   "SDC\DB_SDC_EMS_FLAGS\DB_SDC_EMS_FLAGS.EMS[99]" : Int AT %DB0.DBW0, 1 s
   "SDC\DB_SDC_EMS_FLAGS\DB_SDC_EMS_FLAGS.EMS[100]" : Int AT %DB0.DBW0, 1 s
   "SDC\DB_SDC_EMS_FLAGS\DB_SDC_EMS_FLAGS.EMS[101]" : Int AT %DB0.DBW0, 1 s
   "SDC\DB_SDC_EMS_FLAGS\DB_SDC_EMS_FLAGS.EMS[102]" : Int AT %DB0.DBW0, 1 s
   "SDC\DB_SDC_EMS_FLAGS\DB_SDC_EMS_FLAGS.EMS[103]" : Int AT %DB0.DBW0, 1 s
   "SDC\DB_SDC_EMS_FLAGS\DB_SDC_EMS_FLAGS.EMS[104]" : Int AT %DB0.DBW0, 1 s
   "SDC\DB_SDC_EMS_FLAGS\DB_SDC_EMS_FLAGS.EMS[105]" : Int AT %DB0.DBW0, 1 s
   "SDC\DB_SDC_EMS_FLAGS\DB_SDC_EMS_FLAGS.EMS[106]" : Int AT %DB0.DBW0, 1 s
   "SDC\DB_SDC_EMS_FLAGS\DB_SDC_EMS_FLAGS.EMS[107]" : Int AT %DB0.DBW0, 1 s
   "SDC\DB_SDC_EMS_FLAGS\DB_SDC_EMS_FLAGS.EMS[108]" : Int AT %DB0.DBW0, 1 s
   "SDC\DB_SDC_EMS_FLAGS\DB_SDC_EMS_FLAGS.EMS[109]" : Int AT %DB0.DBW0, 1 s
   "SDC\DB_SDC_EMS_FLAGS\_EMS_Flags_Byte_EMS001" : Int, internal
   "SDC\DB_SDC_EMS_FLAGS\_EMS_Flags_Byte_EMS002" : Int, internal
   "SDC\DB_SDC_EMS_FLAGS\_EMS_Flags_Byte_EMS003" : Int, internal
   "SDC\DB_SDC_EMS_FLAGS\_EMS_Flags_Byte_EMS004" : Int, internal
   "SDC\DB_SDC_EMS_FLAGS\_EMS_Flags_Byte_EMS005" : Int, internal
   "SDC\DB_SDC_EMS_FLAGS\_EMS_Flags_Byte_EMS006" : Int, internal
   "SDC\DB_SDC_EMS_FLAGS\_EMS_Flags_Byte_EMS007" : Int, internal
   "SDC\DB_SDC_EMS_FLAGS\_EMS_Flags_Byte_EMS008" : Int, internal
   "SDC\DB_SDC_EMS_FLAGS\_EMS_Flags_Byte_EMS009" : Int, internal
   "SDC\DB_SDC_EMS_FLAGS\_EMS_Flags_Byte_EMS010" : Int, internal
   "SDC\DB_SDC_EMS_FLAGS\_EMS_Flags_Byte_EMS011" : Int, internal
   "SDC\DB_SDC_EMS_FLAGS\_EMS_Flags_Byte_EMS012" : Int, internal
   "SDC\DB_SDC_EMS_FLAGS\_EMS_Flags_Byte_EMS013" : Int, internal
   "SDC\DB_SDC_EMS_FLAGS\_EMS_Flags_Byte_EMS014" : Int, internal
   "SDC\DB_SDC_EMS_FLAGS\_EMS_Flags_Byte_EMS015" : Int, internal
   "SDC\DB_SDC_EMS_FLAGS\_EMS_Flags_Byte_EMS016" : Int, internal
   "SDC\DB_SDC_EMS_FLAGS\_EMS_Flags_Byte_EMS017" : Int, internal
   "SDC\DB_SDC_EMS_FLAGS\_EMS_Flags_Byte_EMS018" : Int, internal
   "SDC\DB_SDC_EMS_FLAGS\_EMS_Flags_Byte_EMS019" : Int, internal
   "SDC\DB_SDC_EMS_FLAGS\_EMS_Flags_Byte_EMS020" : Int, internal
   "SDC\DB_SDC_EMS_FLAGS\_EMS_Flags_Byte_EMS021" : Int, internal
   "SDC\DB_SDC_EMS_FLAGS\_EMS_Flags_Byte_EMS022" : Int, internal
   "SDC\DB_SDC_EMS_FLAGS\_EMS_Flags_Byte_EMS023" : Int, internal
   "SDC\DB_SDC_EMS_FLAGS\_EMS_Flags_Byte_EMS024" : Int, internal
   "SDC\DB_SDC_EMS_FLAGS\_EMS_Flags_Byte_EMS025" : Int, internal
   "SDC\DB_SDC_EMS_FLAGS\_EMS_Flags_Byte_EMS026" : Int, internal
   "SDC\DB_SDC_EMS_FLAGS\_EMS_Flags_Byte_EMS027" : Int, internal
   "SDC\DB_SDC_EMS_FLAGS\_EMS_Flags_Byte_EMS028" : Int, internal
   "SDC\DB_SDC_EMS_FLAGS\_EMS_Flags_Byte_EMS029" : Int, internal
   "SDC\DB_SDC_EMS_FLAGS\_EMS_Flags_Byte_EMS030" : Int, internal
   "SDC\DB_SDC_EMS_FLAGS\_EMS_Flags_Byte_EMS031" : Int, internal
   "SDC\DB_SDC_EMS_FLAGS\_EMS_Flags_Byte_EMS032" : Int, internal
   "SDC\DB_SDC_EMS_FLAGS\_EMS_Flags_Byte_EMS033" : Int, internal
   "SDC\DB_SDC_EMS_FLAGS\_EMS_Flags_Byte_EMS034" : Int, internal
   "SDC\DB_SDC_EMS_FLAGS\_EMS_Flags_Byte_EMS035" : Int, internal
   "SDC\DB_SDC_EMS_FLAGS\_EMS_Flags_Byte_EMS036" : Int, internal
   "SDC\DB_SDC_EMS_FLAGS\_EMS_Flags_Byte_EMS037" : Int, internal
   "SDC\DB_SDC_EMS_FLAGS\_EMS_Flags_Byte_EMS038" : Int, internal
   "SDC\DB_SDC_EMS_FLAGS\_EMS_Flags_Byte_EMS039" : Int, internal
   "SDC\DB_SDC_EMS_FLAGS\_EMS_Flags_Byte_EMS040" : Int, internal
   "SDC\DB_SDC_EMS_FLAGS\_EMS_Flags_Byte_EMS041" : Int, internal
   "SDC\DB_SDC_EMS_FLAGS\_EMS_Flags_Byte_EMS042" : Int, internal
   "SDC\DB_SDC_EMS_FLAGS\_EMS_Flags_Byte_EMS043" : Int, internal
   "SDC\DB_SDC_EMS_FLAGS\_EMS_Flags_Byte_EMS044" : Int, internal
   "SDC\DB_SDC_EMS_FLAGS\_EMS_Flags_Byte_EMS045" : Int, internal
   "SDC\DB_SDC_EMS_FLAGS\_EMS_Flags_Byte_EMS046" : Int, internal
   "SDC\DB_SDC_EMS_FLAGS\_EMS_Flags_Byte_EMS047" : Int, internal
   "SDC\DB_SDC_EMS_FLAGS\_EMS_Flags_Byte_EMS048" : Int, internal
   "SDC\DB_SDC_EMS_FLAGS\_EMS_Flags_Byte_EMS049" : Int, internal
   "SDC\DB_SDC_EMS_FLAGS\_EMS_Flags_Byte_EMS050" : Int, internal
   "SDC\DB_SDC_EMS_FLAGS\_EMS_Flags_Byte_EMS051" : Int, internal
   "SDC\DB_SDC_EMS_FLAGS\_EMS_Flags_Byte_EMS052" : Int, internal
   "SDC\DB_SDC_EMS_FLAGS\_EMS_Flags_Byte_EMS053" : Int, internal
   "SDC\DB_SDC_EMS_FLAGS\_EMS_Flags_Byte_EMS054" : Int, internal
   "SDC\DB_SDC_EMS_FLAGS\_EMS_Flags_Byte_EMS055" : Int, internal
   "SDC\DB_SDC_EMS_FLAGS\_EMS_Flags_Byte_EMS056" : Int, internal
   "SDC\DB_SDC_EMS_FLAGS\_EMS_Flags_Byte_EMS057" : Int, internal
   "SDC\DB_SDC_EMS_FLAGS\_EMS_Flags_Byte_EMS058" : Int, internal
   "SDC\DB_SDC_EMS_FLAGS\_EMS_Flags_Byte_EMS059" : Int, internal
   "SDC\DB_SDC_EMS_FLAGS\_EMS_Flags_Byte_EMS060" : Int, internal
   "SDC\DB_SDC_EMS_FLAGS\_EMS_Flags_Byte_EMS061" : Int, internal
   "SDC\DB_SDC_EMS_FLAGS\_EMS_Flags_Byte_EMS062" : Int, internal
   "SDC\DB_SDC_EMS_FLAGS\_EMS_Flags_Byte_EMS063" : Int, internal
   "SDC\DB_SDC_EMS_FLAGS\_EMS_Flags_Byte_EMS064" : Int, internal
   "SDC\DB_SDC_EMS_FLAGS\_EMS_Flags_Byte_EMS065" : Int, internal
   "SDC\DB_SDC_EMS_FLAGS\_EMS_Flags_Byte_EMS066" : Int, internal
   "SDC\DB_SDC_EMS_FLAGS\_EMS_Flags_Byte_EMS067" : Int, internal
   "SDC\DB_SDC_EMS_FLAGS\_EMS_Flags_Byte_EMS068" : Int, internal
   "SDC\DB_SDC_EMS_FLAGS\_EMS_Flags_Byte_EMS069" : Int, internal
   "SDC\DB_SDC_EMS_FLAGS\_EMS_Flags_Byte_EMS070" : Int, internal
   "SDC\DB_SDC_EMS_FLAGS\_EMS_Flags_Byte_EMS071" : Int, internal
   "SDC\DB_SDC_EMS_FLAGS\_EMS_Flags_Byte_EMS072" : Int, internal
   "SDC\DB_SDC_EMS_FLAGS\_EMS_Flags_Byte_EMS073" : Int, internal
   "SDC\DB_SDC_EMS_FLAGS\_EMS_Flags_Byte_EMS074" : Int, internal
   "SDC\DB_SDC_EMS_FLAGS\_EMS_Flags_Byte_EMS075" : Int, internal
   "SDC\DB_SDC_EMS_FLAGS\_EMS_Flags_Byte_EMS076" : Int, internal
   "SDC\DB_SDC_EMS_FLAGS\_EMS_Flags_Byte_EMS077" : Int, internal
   "SDC\DB_SDC_EMS_FLAGS\_EMS_Flags_Byte_EMS078" : Int, internal
   "SDC\DB_SDC_EMS_FLAGS\_EMS_Flags_Byte_EMS079" : Int, internal
   "SDC\DB_SDC_EMS_FLAGS\_EMS_Flags_Byte_EMS080" : Int, internal
   "SDC\DB_SDC_EMS_FLAGS\_EMS_Flags_Byte_EMS081" : Int, internal
   "SDC\DB_SDC_EMS_FLAGS\_EMS_Flags_Byte_EMS082" : Int, internal
   "SDC\DB_SDC_EMS_FLAGS\_EMS_Flags_Byte_EMS083" : Int, internal
   "SDC\DB_SDC_EMS_FLAGS\_EMS_Flags_Byte_EMS084" : Int, internal
   "SDC\DB_SDC_EMS_FLAGS\_EMS_Flags_Byte_EMS085" : Int, internal
   "SDC\DB_SDC_EMS_FLAGS\_EMS_Flags_Byte_EMS086" : Int, internal
   "SDC\DB_SDC_EMS_FLAGS\_EMS_Flags_Byte_EMS087" : Int, internal
   "SDC\DB_SDC_EMS_FLAGS\_EMS_Flags_Byte_EMS088" : Int, internal
   "SDC\DB_SDC_EMS_FLAGS\_EMS_Flags_Byte_EMS089" : Int, internal
   "SDC\DB_SDC_EMS_FLAGS\_EMS_Flags_Byte_EMS090" : Int, internal
   "SDC\DB_SDC_EMS_FLAGS\_EMS_Flags_Byte_EMS091" : Int, internal
   "SDC\DB_SDC_EMS_FLAGS\_EMS_Flags_Byte_EMS092" : Int, internal
   "SDC\DB_SDC_EMS_FLAGS\_EMS_Flags_Byte_EMS093" : Int, internal
   "SDC\DB_SDC_EMS_FLAGS\_EMS_Flags_Byte_EMS094" : Int, internal
   "SDC\DB_SDC_EMS_FLAGS\_EMS_Flags_Byte_EMS095" : Int, internal
   "SDC\DB_SDC_EMS_FLAGS\_EMS_Flags_Byte_EMS096" : Int, internal
   "SDC\DB_SDC_EMS_FLAGS\_EMS_Flags_Byte_EMS097" : Int, internal
   "SDC\DB_SDC_EMS_FLAGS\_EMS_Flags_Byte_EMS098" : Int, internal
   "SDC\DB_SDC_EMS_FLAGS\_EMS_Flags_Byte_EMS099" : Int, internal
   "SDC\DB_SDC_EMS_FLAGS\_EMS_Flags_Byte_EMS100" : Int, internal
   "SDC\DB_SDC_EMS_FLAGS\_EMS_Flags_Byte_EMS101" : Int, internal
   "SDC\DB_SDC_EMS_FLAGS\_EMS_Flags_Byte_EMS102" : Int, internal
   "SDC\DB_SDC_EMS_FLAGS\_EMS_Flags_Byte_EMS103" : Int, internal
   "SDC\DB_SDC_EMS_FLAGS\_EMS_Flags_Byte_EMS104" : Int, internal
   "SDC\DB_SDC_EMS_FLAGS\_EMS_Flags_Byte_EMS105" : Int, internal
   "SDC\DB_SDC_EMS_FLAGS\_EMS_Flags_Byte_EMS106" : Int, internal
   "SDC\DB_SDC_EMS_FLAGS\_EMS_Flags_Byte_EMS107" : Int, internal
   "SDC\DB_SDC_EMS_FLAGS\_EMS_Flags_Byte_EMS108" : Int, internal
   "SDC\DB_SDC_EMS_FLAGS\_EMS_Flags_Byte_EMS109" : Int, internal
   "DB_SDC_EMS_FLAGS_HMI_HEADER.DB_NR" : Int = PLC DB_SDC_EMS_FLAGS_HMI.HEADER.DB_NR AT %DB3801.DBW0, 1 s
   "SDC\DB_SDC_EMS_FLAGS\_EMS_Flags_Byte_EMS110" : Int, internal
   "SDC\DB_SDC_EMS_FLAGS\_EMS_Flags_Byte_EMS111" : Int, internal
   "SDC\DB_SDC_EMS_FLAGS\_EMS_Flags_Byte_EMS112" : Int, internal
   "SDC\DB_SDC_EMS_FLAGS\_EMS_Flags_Byte_EMS113" : Int, internal
   "SDC\DB_SDC_EMS_FLAGS\_EMS_Flags_Byte_EMS114" : Int, internal
   "SDC\DB_SDC_EMS_FLAGS\_EMS_Flags_Byte_EMS115" : Int, internal
   "SDC\DB_SDC_EMS_FLAGS\_EMS_Flags_Byte_EMS116" : Int, internal
   "SDC\DB_SDC_EMS_FLAGS\_EMS_Flags_Byte_EMS117" : Int, internal
   "SDC\DB_SDC_EMS_FLAGS\_EMS_Flags_Byte_EMS118" : Int, internal
   "SDC\DB_SDC_EMS_FLAGS\_EMS_Flags_Byte_EMS119" : Int, internal
   "SDC\DB_SDC_EMS_FLAGS\_EMS_Flags_Byte_EMS120" : Int, internal
   "SDC\DB_SDC_EMS_FLAGS\_EMS_Flags_Byte_EMS121" : Int, internal
   "SDC\DB_SDC_EMS_FLAGS\_EMS_Flags_Byte_EMS122" : Int, internal
   "SDC\DB_SDC_EMS_FLAGS\_EMS_Flags_Byte_EMS123" : Int, internal
   "SDC\DB_SDC_EMS_FLAGS\_EMS_Flags_Byte_EMS124" : Int, internal
   "SDC\DB_SDC_EMS_FLAGS\_EMS_Flags_Byte_EMS125" : Int, internal
   "SDC\DB_SDC_EMS_FLAGS\_EMS_Flags_Byte_EMS126" : Int, internal
   "SDC\DB_SDC_EMS_FLAGS\_EMS_Flags_Byte_EMS127" : Int, internal
   "SDC\DB_SDC_EMS_FLAGS\_EMS_Flags_Byte_EMS128" : Int, internal
   "SDC\DB_SDC_EMS_FLAGS\_EMS_Flags_Byte_EMS129" : Int, internal
   "SDC\DB_SDC_EMS_FLAGS\_EMS_Flags_Byte_EMS130" : Int, internal
   "SDC\DB_SDC_EMS_FLAGS\_EMS_Flags_Byte_EMS131" : Int, internal
   "SDC\DB_SDC_EMS_FLAGS\_EMS_Flags_Byte_EMS132" : Int, internal
   "SDC\DB_SDC_EMS_FLAGS\_EMS_Flags_Byte_EMS133" : Int, internal
   "SDC\DB_SDC_EMS_FLAGS\_EMS_Flags_Byte_EMS134" : Int, internal
   "SDC\DB_SDC_EMS_FLAGS\_EMS_Flags_Byte_EMS135" : Int, internal
   "SDC\DB_SDC_EMS_FLAGS\_EMS_Flags_Byte_EMS136" : Int, internal
   "SDC\DB_SDC_EMS_FLAGS\_EMS_Flags_Byte_EMS137" : Int, internal
   "SDC\DB_SDC_EMS_FLAGS\_EMS_Flags_Byte_EMS138" : Int, internal
   "SDC\DB_SDC_EMS_FLAGS\_EMS_Flags_Byte_EMS139" : Int, internal
   "SDC\DB_SDC_EMS_FLAGS\_EMS_Flags_Byte_EMS140" : Int, internal
   "SDC\DB_SDC_EMS_FLAGS\_EMS_Flags_Byte_EMS141" : Int, internal
   "SDC\DB_SDC_EMS_FLAGS\_EMS_Flags_Byte_EMS142" : Int, internal
   "SDC\DB_SDC_EMS_FLAGS\_EMS_Flags_Byte_EMS143" : Int, internal
   "SDC\DB_SDC_EMS_FLAGS\_EMS_Flags_Byte_EMS144" : Int, internal
   "SDC\DB_SDC_EMS_FLAGS\_EMS_Flags_Byte_EMS145" : Int, internal
   "SDC\DB_SDC_EMS_FLAGS\_EMS_Flags_Byte_EMS146" : Int, internal
   "SDC\DB_SDC_EMS_FLAGS\_EMS_Flags_Byte_EMS147" : Int, internal
   "SDC\DB_SDC_EMS_FLAGS\_EMS_Flags_Byte_EMS148" : Int, internal
   "SDC\DB_SDC_EMS_FLAGS\_EMS_Flags_Byte_EMS149" : Int, internal
   "SDC\DB_SDC_EMS_FLAGS\_EMS_Flags_Byte_EMS150" : Int, internal
   "SDC\DB_SDC_EMS_FLAGS\_EMS_Flags_Byte_EMS151" : Int, internal
   "SDC\DB_SDC_EMS_FLAGS\_EMS_Flags_Byte_EMS152" : Int, internal
   "SDC\DB_SDC_EMS_FLAGS\_EMS_Flags_Byte_EMS153" : Int, internal
   "SDC\DB_SDC_EMS_FLAGS\_EMS_Flags_Byte_EMS154" : Int, internal
   "SDC\DB_SDC_EMS_FLAGS\_EMS_Flags_Byte_EMS155" : Int, internal
   "SDC\DB_SDC_EMS_FLAGS\_EMS_Flags_Byte_EMS156" : Int, internal
   "SDC\DB_SDC_EMS_FLAGS\_EMS_Flags_Byte_EMS157" : Int, internal
   "SDC\DB_SDC_EMS_FLAGS\_EMS_Flags_Byte_EMS158" : Int, internal
   "SDC\DB_SDC_EMS_FLAGS\_EMS_Flags_Byte_EMS159" : Int, internal
   "SDC\DB_SDC_EMS_FLAGS\_EMS_Flags_Byte_EMS160" : Int, internal
   "SDC\DB_SDC_EMS_FLAGS\_EMS_Flags_Byte_EMS161" : Int, internal
   "SDC\DB_SDC_EMS_FLAGS\_EMS_Flags_Byte_EMS162" : Int, internal
   "SDC\DB_SDC_EMS_FLAGS\_EMS_Flags_Byte_EMS163" : Int, internal
   "SDC\DB_SDC_EMS_FLAGS\_EMS_Flags_Byte_EMS164" : Int, internal
   "SDC\DB_SDC_EMS_FLAGS\_EMS_Flags_Byte_EMS165" : Int, internal
   "SDC\DB_SDC_EMS_FLAGS\_EMS_Flags_Byte_EMS166" : Int, internal
   "SDC\DB_SDC_EMS_FLAGS\_EMS_Flags_Byte_EMS167" : Int, internal
   "SDC\DB_SDC_EMS_FLAGS\_EMS_Flags_Byte_EMS168" : Int, internal
   "SDC\DB_SDC_EMS_FLAGS\_EMS_Flags_Byte_EMS169" : Int, internal
   "SDC\DB_SDC_EMS_FLAGS\_EMS_Flags_Byte_EMS170" : Int, internal
   "SDC\DB_SDC_EMS_FLAGS\_EMS_Flags_Byte_EMS171" : Int, internal
   "SDC\DB_SDC_EMS_FLAGS\_EMS_Flags_Byte_EMS172" : Int, internal
   "SDC\DB_SDC_EMS_FLAGS\_EMS_Flags_Byte_EMS173" : Int, internal
   "SDC\DB_SDC_EMS_FLAGS\_EMS_Flags_Byte_EMS174" : Int, internal
   "SDC\DB_SDC_EMS_FLAGS\_EMS_Flags_Byte_EMS175" : Int, internal
   "SDC\DB_SDC_EMS_FLAGS\_EMS_Flags_Byte_EMS176" : Int, internal
   "SDC\DB_SDC_EMS_FLAGS\_EMS_Flags_Byte_EMS177" : Int, internal
   "SDC\DB_SDC_EMS_FLAGS\_EMS_Flags_Byte_EMS178" : Int, internal
   "SDC\DB_SDC_EMS_FLAGS\_EMS_Flags_Byte_EMS179" : Int, internal
   "SDC\DB_SDC_EMS_FLAGS\_EMS_Flags_Byte_EMS180" : Int, internal
   "SDC\DB_SDC_EMS_FLAGS\_EMS_Flags_Byte_EMS181" : Int, internal
   "SDC\DB_SDC_EMS_FLAGS\_EMS_Flags_Byte_EMS182" : Int, internal
   "SDC\DB_SDC_EMS_FLAGS\_EMS_Flags_Byte_EMS183" : Int, internal
   "SDC\DB_SDC_EMS_FLAGS\_EMS_Flags_Byte_EMS184" : Int, internal
   "SDC\DB_SDC_EMS_FLAGS\DB_SDC_EMS_FLAGS.EMS[110]" : Int AT %DB0.DBW0, 1 s
   "SDC\DB_SDC_EMS_FLAGS\DB_SDC_EMS_FLAGS.EMS[111]" : Int AT %DB0.DBW0, 1 s
   "SDC\DB_SDC_EMS_FLAGS\DB_SDC_EMS_FLAGS.EMS[112]" : Int AT %DB0.DBW0, 1 s
   "SDC\DB_SDC_EMS_FLAGS\DB_SDC_EMS_FLAGS.EMS[113]" : Int AT %DB0.DBW0, 1 s
   "SDC\DB_SDC_EMS_FLAGS\DB_SDC_EMS_FLAGS.EMS[114]" : Int AT %DB0.DBW0, 1 s
   "SDC\DB_SDC_EMS_FLAGS\DB_SDC_EMS_FLAGS.EMS[115]" : Int AT %DB0.DBW0, 1 s
   "SDC\DB_SDC_EMS_FLAGS\DB_SDC_EMS_FLAGS.EMS[116]" : Int AT %DB0.DBW0, 1 s
   "SDC\DB_SDC_EMS_FLAGS\DB_SDC_EMS_FLAGS.EMS[117]" : Int AT %DB0.DBW0, 1 s
   "SDC\DB_SDC_EMS_FLAGS\DB_SDC_EMS_FLAGS.EMS[118]" : Int AT %DB0.DBW0, 1 s
   "SDC\DB_SDC_EMS_FLAGS\DB_SDC_EMS_FLAGS.EMS[119]" : Int AT %DB0.DBW0, 1 s
   "SDC\DB_SDC_EMS_FLAGS\DB_SDC_EMS_FLAGS.EMS[120]" : Int AT %DB0.DBW0, 1 s
   "SDC\DB_SDC_EMS_FLAGS\DB_SDC_EMS_FLAGS.EMS[121]" : Int AT %DB0.DBW0, 1 s
   "SDC\DB_SDC_EMS_FLAGS\DB_SDC_EMS_FLAGS.EMS[122]" : Int AT %DB0.DBW0, 1 s
   "SDC\DB_SDC_EMS_FLAGS\DB_SDC_EMS_FLAGS.EMS[123]" : Int AT %DB0.DBW0, 1 s
   "SDC\DB_SDC_EMS_FLAGS\DB_SDC_EMS_FLAGS.EMS[124]" : Int AT %DB0.DBW0, 1 s
   "SDC\DB_SDC_EMS_FLAGS\DB_SDC_EMS_FLAGS.EMS[125]" : Int AT %DB0.DBW0, 1 s
   "SDC\DB_SDC_EMS_FLAGS\DB_SDC_EMS_FLAGS.EMS[126]" : Int AT %DB0.DBW0, 1 s
   "SDC\DB_SDC_EMS_FLAGS\DB_SDC_EMS_FLAGS.EMS[127]" : Int AT %DB0.DBW0, 1 s
   "SDC\DB_SDC_EMS_FLAGS\DB_SDC_EMS_FLAGS.EMS[128]" : Int AT %DB0.DBW0, 1 s
   "SDC\DB_SDC_EMS_FLAGS\DB_SDC_EMS_FLAGS.EMS[129]" : Int AT %DB0.DBW0, 1 s
   "SDC\DB_SDC_EMS_FLAGS\DB_SDC_EMS_FLAGS.EMS[130]" : Int AT %DB0.DBW0, 1 s
   "SDC\DB_SDC_EMS_FLAGS\DB_SDC_EMS_FLAGS.EMS[131]" : Int AT %DB0.DBW0, 1 s
   "SDC\DB_SDC_EMS_FLAGS\DB_SDC_EMS_FLAGS.EMS[132]" : Int AT %DB0.DBW0, 1 s
   "SDC\DB_SDC_EMS_FLAGS\DB_SDC_EMS_FLAGS.EMS[133]" : Int AT %DB0.DBW0, 1 s
   "SDC\DB_SDC_EMS_FLAGS\DB_SDC_EMS_FLAGS.EMS[134]" : Int AT %DB0.DBW0, 1 s
   "SDC\DB_SDC_EMS_FLAGS\DB_SDC_EMS_FLAGS.EMS[135]" : Int AT %DB0.DBW0, 1 s
   "SDC\DB_SDC_EMS_FLAGS\DB_SDC_EMS_FLAGS.EMS[136]" : Int AT %DB0.DBW0, 1 s
   "SDC\DB_SDC_EMS_FLAGS\DB_SDC_EMS_FLAGS.EMS[137]" : Int AT %DB0.DBW0, 1 s
   "SDC\DB_SDC_EMS_FLAGS\DB_SDC_EMS_FLAGS.EMS[138]" : Int AT %DB0.DBW0, 1 s
   "SDC\DB_SDC_EMS_FLAGS\DB_SDC_EMS_FLAGS.EMS[139]" : Int AT %DB0.DBW0, 1 s
   "SDC\DB_SDC_EMS_FLAGS\DB_SDC_EMS_FLAGS.EMS[140]" : Int AT %DB0.DBW0, 1 s
   "SDC\DB_SDC_EMS_FLAGS\DB_SDC_EMS_FLAGS.EMS[141]" : Int AT %DB0.DBW0, 1 s
   "SDC\DB_SDC_EMS_FLAGS\DB_SDC_EMS_FLAGS.EMS[142]" : Int AT %DB0.DBW0, 1 s
   "SDC\DB_SDC_EMS_FLAGS\DB_SDC_EMS_FLAGS.EMS[143]" : Int AT %DB0.DBW0, 1 s
   "SDC\DB_SDC_EMS_FLAGS\DB_SDC_EMS_FLAGS.EMS[144]" : Int AT %DB0.DBW0, 1 s
   "SDC\DB_SDC_EMS_FLAGS\DB_SDC_EMS_FLAGS.EMS[145]" : Int AT %DB0.DBW0, 1 s
   "SDC\DB_SDC_EMS_FLAGS\DB_SDC_EMS_FLAGS.EMS[146]" : Int AT %DB0.DBW0, 1 s
   "SDC\DB_SDC_EMS_FLAGS\DB_SDC_EMS_FLAGS.EMS[147]" : Int AT %DB0.DBW0, 1 s
   "SDC\DB_SDC_EMS_FLAGS\DB_SDC_EMS_FLAGS.EMS[148]" : Int AT %DB0.DBW0, 1 s
   "SDC\DB_SDC_EMS_FLAGS\DB_SDC_EMS_FLAGS.EMS[149]" : Int AT %DB0.DBW0, 1 s
   "SDC\DB_SDC_EMS_FLAGS\DB_SDC_EMS_FLAGS.EMS[150]" : Int AT %DB0.DBW0, 1 s
   "SDC\DB_SDC_EMS_FLAGS\DB_SDC_EMS_FLAGS.EMS[151]" : Int AT %DB0.DBW0, 1 s
   "SDC\DB_SDC_EMS_FLAGS\DB_SDC_EMS_FLAGS.EMS[152]" : Int AT %DB0.DBW0, 1 s
   "SDC\DB_SDC_EMS_FLAGS\DB_SDC_EMS_FLAGS.EMS[153]" : Int AT %DB0.DBW0, 1 s
   "SDC\DB_SDC_EMS_FLAGS\DB_SDC_EMS_FLAGS.EMS[154]" : Int AT %DB0.DBW0, 1 s
   "SDC\DB_SDC_EMS_FLAGS\DB_SDC_EMS_FLAGS.EMS[155]" : Int AT %DB0.DBW0, 1 s
   "SDC\DB_SDC_EMS_FLAGS\DB_SDC_EMS_FLAGS.EMS[156]" : Int AT %DB0.DBW0, 1 s
   "SDC\DB_SDC_EMS_FLAGS\DB_SDC_EMS_FLAGS.EMS[157]" : Int AT %DB0.DBW0, 1 s
   "SDC\DB_SDC_EMS_FLAGS\DB_SDC_EMS_FLAGS.EMS[158]" : Int AT %DB0.DBW0, 1 s
   "SDC\DB_SDC_EMS_FLAGS\DB_SDC_EMS_FLAGS.EMS[159]" : Int AT %DB0.DBW0, 1 s
   "SDC\DB_SDC_EMS_FLAGS\DB_SDC_EMS_FLAGS.EMS[160]" : Int AT %DB0.DBW0, 1 s
   "SDC\DB_SDC_EMS_FLAGS\DB_SDC_EMS_FLAGS.EMS[161]" : Int AT %DB0.DBW0, 1 s
   "SDC\DB_SDC_EMS_FLAGS\DB_SDC_EMS_FLAGS.EMS[162]" : Int AT %DB0.DBW0, 1 s
   "SDC\DB_SDC_EMS_FLAGS\DB_SDC_EMS_FLAGS.EMS[163]" : Int AT %DB0.DBW0, 1 s
   "SDC\DB_SDC_EMS_FLAGS\DB_SDC_EMS_FLAGS.EMS[164]" : Int AT %DB0.DBW0, 1 s
   "SDC\DB_SDC_EMS_FLAGS\DB_SDC_EMS_FLAGS.EMS[165]" : Int AT %DB0.DBW0, 1 s
   "SDC\DB_SDC_EMS_FLAGS\DB_SDC_EMS_FLAGS.EMS[166]" : Int AT %DB0.DBW0, 1 s
   "SDC\DB_SDC_EMS_FLAGS\DB_SDC_EMS_FLAGS.EMS[167]" : Int AT %DB0.DBW0, 1 s
   "SDC\DB_SDC_EMS_FLAGS\DB_SDC_EMS_FLAGS.EMS[168]" : Int AT %DB0.DBW0, 1 s
   "SDC\DB_SDC_EMS_FLAGS\DB_SDC_EMS_FLAGS.EMS[169]" : Int AT %DB0.DBW0, 1 s
   "SDC\DB_SDC_EMS_FLAGS\DB_SDC_EMS_FLAGS.EMS[170]" : Int AT %DB0.DBW0, 1 s
   "SDC\DB_SDC_EMS_FLAGS\DB_SDC_EMS_FLAGS.EMS[171]" : Int AT %DB0.DBW0, 1 s
   "SDC\DB_SDC_EMS_FLAGS\DB_SDC_EMS_FLAGS.EMS[172]" : Int AT %DB0.DBW0, 1 s
   "SDC\DB_SDC_EMS_FLAGS\DB_SDC_EMS_FLAGS.EMS[173]" : Int AT %DB0.DBW0, 1 s
   "SDC\DB_SDC_EMS_FLAGS\DB_SDC_EMS_FLAGS.EMS[174]" : Int AT %DB0.DBW0, 1 s
   "SDC\DB_SDC_EMS_FLAGS\DB_SDC_EMS_FLAGS.EMS[175]" : Int AT %DB0.DBW0, 1 s
   "SDC\DB_SDC_EMS_FLAGS\DB_SDC_EMS_FLAGS.EMS[176]" : Int AT %DB0.DBW0, 1 s
   "SDC\DB_SDC_EMS_FLAGS\DB_SDC_EMS_FLAGS.EMS[177]" : Int AT %DB0.DBW0, 1 s
   "SDC\DB_SDC_EMS_FLAGS\DB_SDC_EMS_FLAGS.EMS[178]" : Int AT %DB0.DBW0, 1 s
   "SDC\DB_SDC_EMS_FLAGS\DB_SDC_EMS_FLAGS.EMS[179]" : Int AT %DB0.DBW0, 1 s
   "SDC\DB_SDC_EMS_FLAGS\DB_SDC_EMS_FLAGS.EMS[180]" : Int AT %DB0.DBW0, 1 s
   "SDC\DB_SDC_EMS_FLAGS\DB_SDC_EMS_FLAGS.EMS[181]" : Int AT %DB0.DBW0, 1 s
   "SDC\DB_SDC_EMS_FLAGS\DB_SDC_EMS_FLAGS.EMS[182]" : Int AT %DB0.DBW0, 1 s
   "SDC\DB_SDC_EMS_FLAGS\DB_SDC_EMS_FLAGS.EMS[183]" : Int AT %DB0.DBW0, 1 s
   "SDC\DB_SDC_EMS_FLAGS\DB_SDC_EMS_FLAGS.EMS[184]" : Int AT %DB0.DBW0, 1 s

HMI tags "DB_SDC_EMS"
   "SDC\DB_SDC_EMS\EMS[XXX].DISTANCE" : DInt AT %DB0.DBD0, 1 s   // Abstand zum vorangehenden EMS / distance to preciding EMS
   "SDC\DB_SDC_EMS\_Byte_EMS[XXX].ABS_POS" : Int, internal   // Absolute Position / absolute Positon
   "SDC\DB_SDC_EMS\EMS[XXX].IF_I_EMS.STAT" : DWord AT %DB0.DBD0, 1 s
   "SDC\DB_SDC_EMS\EMS[XXX].PRECEDING_EMS" : Int AT %DB0.DBW0, 1 s   // preciding EMS
   "SDC\DB_SDC_EMS\_Byte_EMS[XXX].TS_STAT.VAL.SEK" : Int, internal   // Sektion
   "SDC\DB_SDC_EMS\_Byte_EMS[XXX].DISTANCE" : Int, internal   // Abstand zum vorangehenden EMS / distance to preciding EMS
   "DB_SDC_EMS_HMI_HEADER.START_HMI" : Int = PLC DB_SDC_EMS_HMI.HEADER.START_HMI AT %DB3814.DBW16, 1 s   // Startadresse HMI
   "SDC\DB_SDC_EMS\EMS[XXX].IF_I_EMS.EA1" : DWord AT %DB0.DBD0, 1 s
   "SDC\DB_SDC_EMS\HMI[XX].PROFIL_Nr" : Int AT %DB0.DBW0, 1 s   // Profilnummer
   "SDC\DB_SDC_EMS\_EMS_HMI_Byte_16" : Int, internal
   "SDC\DB_SDC_EMS\HMI[XX].T_EDIT" : Bool AT %DB0.DBX0.0, 1 s   // Taster Editieren für Pult aktivieren
   "SDC\DB_SDC_EMS\_EMS_HMI_Byte_18" : Int, internal
   "SDC\DB_SDC_EMS\EMS[XXX].FKT_RESET" : Word AT %DB0.DBW0, 1 s   // EMS zur Reperatur / EMS to Repair
   "SDC\DB_SDC_EMS\EMS[XXX].IF_Q_EMS.D_SETSPEED" : DInt AT %DB0.DBD0, 1 s   // set value: drive speed (mm/min)
   "SDC\DB_SDC_EMS\_Byte_EMS[XXX].CYCLE_COUNTER" : Int, internal   // Zykluszähler / Cycle Counter
   "SDC\DB_SDC_EMS\HMI[XX].FR_EDIT" : Bool AT %DB0.DBX0.0, 1 s   // Freigabe Editieren
   "SDC\DB_SDC_EMS\_Byte_EMS[XXX].IF_I_EMS.H_POS" : Int, internal
   "SDC\DB_SDC_EMS\EMS[XXX].TS_STAT.SERIES" : Array [0..3] of Char AT %DB0.DBX0.0, 1 s   // Entwicklungs Serie Karosse (e.g. E-90, E-87 ) / Development series body (e.g. E-90, E-87 )
   "SDC\DB_SDC_EMS\EMS[XXX].IF_Q_EMS.D_SETPOS" : DInt AT %DB0.DBD0, 1 s   // Setpoint: drive position in mm
   "SDC\DB_SDC_EMS\HMI[XX].BILD_Nr_Alt" : Int AT %DB0.DBW0, 1 s   // Bild_Nr alt
   "SDC\DB_SDC_EMS\EMS[XXX].IF_Q_EMS.H_SETSPEED" : Int AT %DB0.DBW0, 1 s   // Setpoint: hoist speed (mm/min)
   "SDC\DB_SDC_EMS\_EMS_HMI_Byte_10" : Int, internal
   "SDC\DB_SDC_EMS\EMS[XXX].IF_I_EMS.H_POS" : Int AT %DB0.DBW0, 1 s
   "SDC\DB_SDC_EMS\_Byte_EMS[XXX].IF_Q_EMS.D_SETPOS" : Int, internal   // Setpoint: drive position in mm Pointer
   "SDC\DB_SDC_EMS\HMI[XX].EMS_Nr" : Int AT %DB0.DBW0, 1 s   // Sektionsnummer
   "SDC\DB_SDC_EMS\_Byte_EMS[XXX].PRECEDING_EMS" : Int, internal   // preciding EMS
   "SDC\DB_SDC_EMS\_Byte_EMS[XXX].IF_I_EMS.STAT" : Int, internal
   "SDC\DB_SDC_EMS\_EMS_HMI_Byte_09" : Int, internal
   "SDC\DB_SDC_EMS\_Byte_EMS[XXX].ERRORS_SDC" : Int, internal   // Fehler SDC Pointer / Faults SDC Pointer
   "SDC\DB_SDC_EMS\EMS[XXX].FLAGS" : Word AT %DB0.DBW0, 1 s   // EMS antrieb vorhanden / EMSdriver present
   "SDC\DB_SDC_EMS\_Byte_EMS[XXX].IF_I_EMS.EA2" : Int, internal
   "SDC\DB_SDC_EMS\EMS[XXX].ERRORS_SDC" : Word AT %DB0.DBW0, 1 s   // Fehler SDC / Faults SDC
   "SDC\DB_SDC_EMS\HMI[XX].T_SAVE" : Bool AT %DB0.DBX0.2, 1 s   // Taster speichern
   "SDC\DB_SDC_EMS\_Byte_EMS[XXX].PROFIL" : Int, internal   // Profile Number
   "SDC\DB_SDC_EMS\_Byte_EMS[XXX].FLAGS" : Int, internal   // EMS antrieb vorhanden / EMSdriver present
   "DB_SDC_EMS_1_HEADER.START_EMS" : Int = PLC DB_SDC_EMS_1.HEADER.START_EMS AT %DB3714.DBW6, 1 s   // Startadresse der EMS Daten im Daten DB
   "SDC\DB_SDC_EMS\EMS[XXX].IF_I_EMS.EA2" : DWord AT %DB0.DBD0, 1 s
   "SDC\DB_SDC_EMS\EMS[XXX].TS_STAT.VAL.SEK" : Int AT %DB0.DBW0, 1 s   // Sektion
      on ChangeValue: "SDC_TS_REFERENCE"("SDC\DB_SDC_EMS\EMS[XXX].TS_STAT.VAL.SEK")
   "SDC\DB_SDC_EMS\EMS[XXX].IF_I_EMS.D_POS" : DInt AT %DB0.DBD0, 1 s
   "SDC\DB_SDC_EMS\_Byte_EMS[XXX].IF_Q_EMS.H_SETSPEED" : Int, internal   // Setpoint: hoist speed (mm/min) Pointer
   "DB_SDC_EMS_1_HEADER.LAENGE_EMS" : Int = PLC DB_SDC_EMS_1.HEADER.LAENGE_EMS AT %DB3714.DBW8, 1 s   // Länge Eingänge pro EMS
   "SDC\DB_SDC_EMS\_EMS_HMI_Byte_19" : Int, internal
   "DB_SDC_EMS_1_HEADER.MIN_NR_EMS" : Int = PLC DB_SDC_EMS_1.HEADER.MIN_NR_EMS AT %DB3714.DBW2, 1 s   // Niedrigste EMS Nummer im Daten DB
   "SDC\DB_SDC_EMS\_Byte_EMS[XXX].IF_Q_EMS.H_SETPOS" : Int, internal   // Setpoint: hoist position (mm) Pointer
   "SDC\DB_SDC_EMS\_Byte_EMS[XXX].IF_I_EMS.EA1" : Int, internal
   "SDC\DB_SDC_EMS\_Intern_DB_EMS_Nr" : Int, internal
   "SDC\DB_SDC_EMS\HMI[XX].ER_DATA" : Bool AT %DB0.DBX0.1, 1 s   // Daten Fehlerhaft
   "DB_SDC_EMS_1_HEADER.OFFSET_EMS_FKT" : Int = PLC DB_SDC_EMS_1.HEADER.OFFSET_EMS_FKT AT %DB3714.DBW14, 1 s   // Offset EMS Funktions
   "SDC\DB_SDC_EMS\EMS[XXX].IF_Q_EMS.H_SETPOS" : Int AT %DB0.DBW0, 1 s   // Setpoint: hoist position (mm)
   "SDC\DB_SDC_EMS\_Byte_EMS[XXX].IF_I_EMS.ERROR" : Int, internal   // Fehlernummer Pointer / Error number Pointer
   "SDC\DB_SDC_EMS\_Byte_EMS[XXX].FKT_RESET" : Int, internal   // EMS zur Reperatur / EMS to Repair
   "SDC\DB_SDC_EMS\EMS[XXX].IF_Q_EMS.CONT" : DWord AT %DB0.DBD0, 1 s
   "DB_SDC_EMS_HMI_HEADER.OFFEST_HMI_DATA" : Int = PLC DB_SDC_EMS_HMI.HEADER.OFFEST_HMI_DATA AT %DB3814.DBW18, 1 s   // Offestadresse der HMI EMS Data
   "SDC\DB_SDC_EMS\_Byte_EMS[XXX].FKT_SET" : Int, internal   // EMS zur Reperatur / EMS to Repair
   "SDC\DB_SDC_EMS\HMI[XX].PULT_Nr_EDIT" : Int AT %DB0.DBW0, 1 s   // Pult Nr Editieren Aktiv (HMI 1 = Master)
   "SDC\DB_SDC_EMS\_EMS_HMI_Byte_00" : Int, internal
   "DB_SDC_EMS_1_HEADER.MAX_NR_EMS" : Int = PLC DB_SDC_EMS_1.HEADER.MAX_NR_EMS AT %DB3714.DBW4, 1 s   // Höchste EMS Nummer im Daten DB
   "SDC\DB_SDC_EMS\EMS[XXX].IF_I_EMS.ERROR" : Int AT %DB0.DBW0, 1 s   // Fehlernummer / Error number
   "DB_SDC_EMS_1_HEADER.OFFSET_EMS_SEK_STAT" : Int = PLC DB_SDC_EMS_1.HEADER.OFFSET_EMS_SEK_STAT AT %DB3714.DBW10, 1 s   // Offset EMS Data
   "DB_SDC_EMS_1_HEADER.LAENGE_EMS_SEK_STAT" : Int = PLC DB_SDC_EMS_1.HEADER.LAENGE_EMS_SEK_STAT AT %DB3714.DBW12, 1 s   // Länge EMS Data
   "SDC\DB_SDC_EMS\_Byte_EMS[XXX].TS_STAT.SERIES" : Int, internal   // Entwicklungs Serie Karosse (e.g. E-90, E-87 ) / Development series body (e.g. E-90, E-87 )
   "SDC\DB_SDC_EMS\HMI[XX].BILD_Nr" : Int AT %DB0.DBW0, 1 s   // Bild_Nr aktiv
   "SDC\DB_SDC_EMS\EMS[XXX].CYCLE_COUNTER" : Int AT %DB0.DBW0, 1 s   // Zykluszähler / Cycle Counter
   "SDC\DB_SDC_EMS\EMS[XXX].FKT_SET" : Word AT %DB0.DBW0, 1 s   // EMS zur Reperatur / EMS to Repair
      on ChangeValue: ResetBit("SDC\DB_SDC_EMS\_Intern_EMS_FKT_Info_Rep_1_on"); ResetBit("SDC\DB_SDC_EMS\_Intern_EMS_FKT_Info_Rep_2_on")
   "SDC\DB_SDC_EMS\HMI[XX].T_LOAD" : Bool AT %DB0.DBX0.3, 1 s   // Taster laden
   "SDC\DB_SDC_EMS\_EMS_HMI_Byte_12" : Int, internal
   "SDC\DB_SDC_EMS\_EMS_HMI_Byte_04" : Int, internal
   "DB_SDC_EMS_HMI_HMI[1].PULT_Nr_EDIT" : Int = PLC DB_SDC_EMS_HMI.HMI[1].PULT_Nr_EDIT AT %DB3814.DBW20, 1 s   // Pult Nr Editieren Aktiv (HMI 1 = Master)
   "SDC\DB_SDC_EMS\_EMS_HMI_Byte_14" : Int, internal
   "SDC\DB_SDC_EMS\_EMS_HMI_Byte_06" : Int, internal
   "SDC\DB_SDC_EMS\_Byte_EMS[XXX].IF_I_EMS.D_POS" : Int, internal
   "SDC\DB_SDC_EMS\_EMS_HMI_Byte_08" : Int, internal
   "SDC\DB_SDC_EMS\EMS[XXX].PROFIL" : Int AT %DB0.DBW0, 1 s   // Profile Number
      on ChangeValue: "SDC_GLOBAL_REFERENCE_PROFIL"("SDC\DB_SDC_EMS\EMS[XXX].PROFIL")
   "SDC\DB_SDC_EMS\_EMS_HMI_Byte_02" : Int, internal
   "SDC\DB_SDC_EMS\EMS[XXX].ABS_POS" : DInt AT %DB0.DBD0, 1 s   // absolute Positon
   "SDC\DB_SDC_EMS\HMI[XX].T_RESET_BED" : Bool AT %DB0.DBX0.1, 1 s   // Taster Reset Bedienfreigabe Pult Nr Bedienung
   "SDC\DB_SDC_EMS\_Byte_EMS[XXX].IF_Q_EMS.CONT" : Int, internal
   "SDC\DB_SDC_EMS\_Byte_EMS[XXX].IF_Q_EMS.D_SETSPEED" : Int, internal   // set value: drive speed (mm/min) Pointer
   "SDC\DB_SDC_EMS\_Byte_EMS[XXX].TS_STAT.VAL.ERROR" : Int, internal   // Sektion
   "SDC\DB_SDC_EMS\EMS[XXX].TS_STAT.VAL.ERROR" : Int AT %DB0.DBW0, 1 s   // Sektion
      on ChangeValue: SetTag("_DB_SDC_ERRORS.Error_nr", "SDC\DB_SDC_EMS\EMS[XXX].TS_STAT.VAL.ERROR")
   "DB_SDC_EMS_HMI_HEADER.DB_NR" : Int = PLC DB_SDC_EMS_HMI.HEADER.DB_NR AT %DB3814.DBW0, 1 s   // DB Nummer
   "SDC\DB_SDC_EMS\_Byte_EMS[XXX].IF_Q_EMS.T_SETPOS" : Int, internal   // Setpoint: hoist position (mm) Pointer
   "SDC\DB_SDC_EMS\_Byte_EMS[XXX].IF_Q_EMS.T_SETSPEED" : Int, internal   // Setpoint: hoist speed (mm/min) Pointer
   "SDC\DB_SDC_EMS\EMS[XXX].IF_Q_EMS.T_SETPOS" : Int AT %DB0.DBW0, 1 s   // Setpoint: hoist position (mm)
   "SDC\DB_SDC_EMS\EMS[XXX].IF_Q_EMS.T_SETSPEED" : Int AT %DB0.DBW0, 1 s   // Setpoint: hoist speed (mm/min)
   "SDC\DB_SDC_EMS\_Byte_EMS[XXX].IF_I_EMS.T_POS" : Int, internal
   "SDC\DB_SDC_EMS\EMS[XXX].IF_I_EMS.T_POS" : Int AT %DB0.DBW0, 1 s
   "SDC\DB_SDC_EMS\_Byte_EMS[XXX].FKT_INFO_REP_1" : Int, internal
   "SDC\DB_SDC_EMS\_Byte_EMS[XXX].FKT_INFO_REP_2" : Int, internal
   "SDC\DB_SDC_EMS\EMS[XXX].FKT_INFO_REP_1" : Int AT %DB0.DBW0, 1 s
   "SDC\DB_SDC_EMS\EMS[XXX].FKT_INFO_REP_2" : Int AT %DB0.DBW0, 1 s
   "SDC\DB_SDC_EMS\_Intern_EMS_FKT_Info_Rep_1_on" : Bool, internal
   "SDC\DB_SDC_EMS\_Intern_EMS_FKT_Info_Rep_2_on" : Bool, internal
   "SDC\DB_SDC_EMS\EMS[XXX].IF_I_EMS.EA3" : Word AT %DB0.DBW0, 1 s
   "SDC\DB_SDC_EMS\_Byte_EMS[XXX].IF_I_EMS.EA3" : Int, internal
   "SDC\DB_SDC_EMS\_Byte_EMS[XXX].VersNo[0]" : Int, internal   // Zykluszähler / Cycle Counter
   "SDC\DB_SDC_EMS\_Byte_EMS[XXX].VersNo[1]" : Int, internal   // Zykluszähler / Cycle Counter
   "SDC\DB_SDC_EMS\EMS[XXX].VersNo[0]" : Byte AT %DB0.DBB0, 1 s   // Zykluszähler / Cycle Counter
   "SDC\DB_SDC_EMS\EMS[XXX].VersNo[1]" : Byte AT %DB0.DBB0, 1 s   // Zykluszähler / Cycle Counter

HMI tags "DB_SDC_SIM"
   "DB_SDC_EMS_SIM_PAR.ON" : Bool = PLC DB_SDC_EMS_SIM.PAR.ON AT %DB3726.DBX40.0, 1 s   // Simulation ON "1"
   "DB_SDC_EMS_SIM_PAR.LEAP_AKT" : Array [0..19] of Bool = PLC DB_SDC_EMS_SIM.PAR.LEAP_AKT AT %DB3726.DBX32.0, 1 s   // Leap Aktiv
   "DB_SDC_EMS_SIM_PAR.BARCODE_START" : DInt = PLC DB_SDC_EMS_SIM.PAR.BARCODE_START AT %DB3726.DBD20, 1 s   // min Barcodevalue
   "DB_SDC_EMS_SIM_PAR.HUB_ENDE" : Int = PLC DB_SDC_EMS_SIM.PAR.HUB_ENDE AT %DB3726.DBW30, 1 s   // max Hoistvalue
   "DB_SDC_EMS_SIM_EMS[2].D_POS" : DInt = PLC DB_SDC_EMS_SIM.EMS[2].D_POS AT %DB3726.DBD90, 1 s   // Antriebsposition in mm / Drive position in mm
   "DB_SDC_EMS_SIM_PAR.BARCODE_ENDE" : DInt = PLC DB_SDC_EMS_SIM.PAR.BARCODE_ENDE AT %DB3726.DBD24, 1 s   // max Barcodevalue
   "DB_SDC_EMS_SIM_PAR.HUB_START" : Int = PLC DB_SDC_EMS_SIM.PAR.HUB_START AT %DB3726.DBW28, 1 s   // min Hoistvalue
   "DB_SDC_EMS_SIM_EMS[1].D_POS" : DInt = PLC DB_SDC_EMS_SIM.EMS[1].D_POS AT %DB3726.DBD50, 1 s   // Antriebsposition in mm / Drive position in mm
   "DB_SDC_EMS_SIM_EMS[3].D_POS" : DInt = PLC DB_SDC_EMS_SIM.EMS[3].D_POS AT %DB3726.DBD130, 1 s   // Antriebsposition in mm / Drive position in mm

HMI tags "DB_SDC_ERRORS"
   "DB_SDC_ERRORS_HEADER.DB_NR" : Int = PLC DB_SDC_ERRORS.HEADER.DB_NR AT %DB3722.DBW0, 1 s
   "DB_SDC_ERRORS_HEADER.MIN_NR_EMS" : Int = PLC DB_SDC_ERRORS.HEADER.MIN_NR_EMS AT %DB3722.DBW2, 1 s
   "DB_SDC_ERRORS_HEADER.MAX_NR_EMS" : Int = PLC DB_SDC_ERRORS.HEADER.MAX_NR_EMS AT %DB3722.DBW4, 1 s
   "DB_SDC_ERRORS_HEADER.START_EMS" : Int = PLC DB_SDC_ERRORS.HEADER.START_EMS AT %DB3722.DBW6, 1 s
   "DB_SDC_ERRORS_HEADER.LAENGE_EMS_StörungS" : Int = PLC DB_SDC_ERRORS.HEADER.LAENGE_EMS_StörungS AT %DB3722.DBW8, 1 s
   "DB_SDC_ERRORS.EMS[XXX].GEN_1" : Word AT %DB0.DBW0, 1 s
   "_Byte_DB_SDC_ERRORS.EMS[XXX].GEN_1" : UInt, internal
   "DB_SDC_ERRORS.EMS[XXX].GEN_2" : Word AT %DB0.DBW0, 1 s
   "_Byte_DB_SDC_ERRORS.EMS[XXX].GEN_2" : UInt, internal
   "DB_SDC_ERRORS.EMS[XXX].GEN_3" : Word AT %DB0.DBW0, 1 s
   "_Byte_DB_SDC_ERRORS.EMS[XXX].GEN_3" : UInt, internal
   "DB_SDC_ERRORS.EMS[XXX].GEN_4" : Word AT %DB0.DBW0, 1 s
   "_Byte_DB_SDC_ERRORS.EMS[XXX].GEN_4" : UInt, internal
   "DB_SDC_ERRORS.EMS[XXX].DRIVE_1" : Word AT %DB0.DBW0, 1 s
   "_Byte_DB_SDC_ERRORS.EMS[XXX].DRIVE_1" : UInt, internal
   "DB_SDC_ERRORS.EMS[XXX].DRIVE_2" : Word AT %DB0.DBW0, 1 s
   "_Byte_DB_SDC_ERRORS.EMS[XXX].DRIVE_2" : UInt, internal
   "DB_SDC_ERRORS.EMS[XXX].FC_DRIVE_1" : Word AT %DB0.DBW0, 1 s
   "_Byte_DB_SDC_ERRORS.EMS[XXX].FC_DRIVE_1" : UInt, internal
   "DB_SDC_ERRORS.EMS[XXX].FC_DRIVE_2" : Word AT %DB0.DBW0, 1 s
   "_Byte_DB_SDC_ERRORS.EMS[XXX].FC_DRIVE_2" : UInt, internal
   "DB_SDC_ERRORS.EMS[XXX].SAFETY_DRIVE" : Word AT %DB0.DBW0, 1 s
   "_Byte_DB_SDC_ERRORS.EMS[XXX].SAFETY_DRIVE" : UInt, internal
   "_Byte_DB_SDC_ERRORS.EMS[XXX].HOIST_1" : UInt, internal
   "DB_SDC_ERRORS.EMS[XXX].HOIST_2" : Word AT %DB0.DBW0, 1 s
   "_Byte_DB_SDC_ERRORS.EMS[XXX].HOIST_2" : UInt, internal
   "DB_SDC_ERRORS.EMS[XXX].FC_HOIST_1" : Word AT %DB0.DBW0, 1 s
   "_Byte_DB_SDC_ERRORS.EMS[XXX].FC_HOIST_1" : UInt, internal
   "DB_SDC_ERRORS.EMS[XXX].FC_HOIST_2" : Word AT %DB0.DBW0, 1 s
   "_Byte_DB_SDC_ERRORS.EMS[XXX].FC_HOIST_2" : UInt, internal
   "DB_SDC_ERRORS.EMS[XXX].SAFETY_HOIST" : Word AT %DB0.DBW0, 1 s
   "_Byte_DB_SDC_ERRORS.EMS[XXX].SAFETY_HOIST" : UInt, internal
   "DB_SDC_ERRORS.EMS[XXX].HOIST_1" : Word AT %DB0.DBW0, 1 s
   "_Byte_DB_SDC_ERRORS.EMS[XXX].TILT_1" : UInt, internal
   "DB_SDC_ERRORS.EMS[XXX].TILT_2" : Word AT %DB0.DBW0, 1 s
   "_Byte_DB_SDC_ERRORS.EMS[XXX].TILT_2" : UInt, internal
   "DB_SDC_ERRORS.EMS[XXX].FC_TILT_1" : Word AT %DB0.DBW0, 1 s
   "_Byte_DB_SDC_ERRORS.EMS[XXX].FC_TILT_1" : UInt, internal
   "DB_SDC_ERRORS.EMS[XXX].FC_TILT_2" : Word AT %DB0.DBW0, 1 s
   "_Byte_DB_SDC_ERRORS.EMS[XXX].FC_TILT_2" : UInt, internal
   "DB_SDC_ERRORS.EMS[XXX].SAFETY_TILT" : Word AT %DB0.DBW0, 1 s
   "_Byte_DB_SDC_ERRORS.EMS[XXX].SAFETY_TILT" : UInt, internal
   "DB_SDC_ERRORS.EMS[XXX].TILT_1" : Word AT %DB0.DBW0, 1 s
   "DB_SDC_ERRORS.EMS[XXX].SDC" : Word AT %DB0.DBW0, 1 s
   "_Byte_DB_SDC_ERRORS.EMS[XXX].SDC" : UInt, internal
   "DB_SDC_ERRORS.SDC" : Word AT %DB3722.DBW20020, 1 s
   "_DB_SDC_ERRORS.Error_nr" : Int, internal
